   "Carrier_55_Carrier_Number_Echo" AT %QW3102 : Word;
   "Carrier_55_Carrier_Position_Echo" AT %QD3104 : DWord;
   "Carrier_55_Next_Carrier_Number" AT %QW3108 : Word;
   "Carrier_55_Next_Stop_Position" AT %QD3110 : DWord;
   "Carrier_55_Drive_Command_Speed" AT %QW3114 : Word;
   "Carrier_55_Duplicate_Carrier_Number" AT %QW3116 : Word;
   "Carrier_55_First_Duplicate_Carrier_Position" AT %QD3118 : DWord;
   "Carrier_55_Second_Duplicate_Carrier_Position" AT %QD3122 : DWord;
   "Carrier_55_CommandWord" AT %QW3126 : Word;
   "Carrier_55_Heartbeat" AT %Q3126.0 : Bool;
   "Carrier_55_Drive_Forward_Command" AT %Q3126.1 : Bool;
   "Carrier_55_Fault_Reset" AT %Q3126.2 : Bool;
   "Carrier_55_At_Command_Position" AT %Q3126.3 : Bool;
   "Carrier_55_Duplicate_Carrier_Fault" AT %Q3126.4 : Bool;
   "Carrier_55_Motion_On_Fault" AT %Q3126.5 : Bool;
   "Carrier_55_Motion_Off_Fault" AT %Q3126.6 : Bool;
   "Carrier_55_Carrier_Spacing_Fault" AT %Q3126.7 : Bool;
   "Carrier_56_Carrier_In_Zone" AT %QW3150 : Word;
   "Carrier_56_Carrier_Number_Echo" AT %QW3152 : Word;
   "Carrier_56_Carrier_Position_Echo" AT %QD3154 : DWord;
   "Carrier_56_Next_Carrier_Number" AT %QW3158 : Word;
   "Carrier_56_Next_Stop_Position" AT %QD3160 : DWord;
   "Carrier_56_Drive_Command_Speed" AT %QW3164 : Word;
   "Carrier_56_Duplicate_Carrier_Number" AT %QW3166 : Word;
   "Carrier_56_First_Duplicate_Carrier_Position" AT %QD3168 : DWord;
   "Carrier_56_Second_Duplicate_Carrier_Position" AT %QD3172 : DWord;
   "Carrier_56_CommandWord" AT %QW3176 : Word;
   "Carrier_56_Heartbeat" AT %Q3176.0 : Bool;
   "Carrier_56_Drive_Forward_Command" AT %Q3176.1 : Bool;
   "Carrier_56_Fault_Reset" AT %Q3176.2 : Bool;
   "Carrier_56_At_Command_Position" AT %Q3176.3 : Bool;
   "Carrier_56_Duplicate_Carrier_Fault" AT %Q3176.4 : Bool;
   "Carrier_56_Motion_On_Fault" AT %Q3176.5 : Bool;
   "Carrier_56_Motion_Off_Fault" AT %Q3176.6 : Bool;
   "Carrier_56_Carrier_Spacing_Fault" AT %Q3176.7 : Bool;
   "Carrier_57_Carrier_In_Zone" AT %QW3200 : Word;
   "Carrier_57_Carrier_Number_Echo" AT %QW3202 : Word;
   "Carrier_57_Carrier_Position_Echo" AT %QD3204 : DWord;
   "Carrier_57_Next_Carrier_Number" AT %QW3208 : Word;
   "Carrier_57_Next_Stop_Position" AT %QD3210 : DWord;
   "Carrier_57_Drive_Command_Speed" AT %QW3214 : Word;
   "Carrier_57_Duplicate_Carrier_Number" AT %QW3216 : Word;
   "Carrier_57_First_Duplicate_Carrier_Position" AT %QD3218 : DWord;
   "Carrier_57_Second_Duplicate_Carrier_Position" AT %QD3222 : DWord;
   "Carrier_57_CommandWord" AT %QW3226 : Word;
   "Carrier_57_Heartbeat" AT %Q3226.0 : Bool;
   "Carrier_57_Drive_Forward_Command" AT %Q3226.1 : Bool;
   "Carrier_57_Fault_Reset" AT %Q3226.2 : Bool;
   "Carrier_57_At_Command_Position" AT %Q3226.3 : Bool;
   "Carrier_57_Duplicate_Carrier_Fault" AT %Q3226.4 : Bool;
   "Carrier_57_Motion_On_Fault" AT %Q3226.5 : Bool;
   "Carrier_57_Motion_Off_Fault" AT %Q3226.6 : Bool;
   "Carrier_57_Carrier_Spacing_Fault" AT %Q3226.7 : Bool;
   "Carrier_58_Carrier_In_Zone" AT %QW3250 : Word;
   "Carrier_58_Carrier_Number_Echo" AT %QW3252 : Word;
   "Carrier_58_Carrier_Position_Echo" AT %QD3254 : DWord;
   "Carrier_58_Next_Carrier_Number" AT %QW3258 : Word;
   "Carrier_58_Next_Stop_Position" AT %QD3260 : DWord;
   "Carrier_58_Drive_Command_Speed" AT %QW3264 : Word;
   "Carrier_58_Duplicate_Carrier_Number" AT %QW3266 : Word;
   "Carrier_58_First_Duplicate_Carrier_Position" AT %QD3268 : DWord;
   "Carrier_58_Second_Duplicate_Carrier_Position" AT %QD3272 : DWord;
   "Carrier_58_CommandWord" AT %QW3276 : Word;
   "Carrier_58_Heartbeat" AT %Q3276.0 : Bool;
   "Carrier_58_Drive_Forward_Command" AT %Q3276.1 : Bool;
   "Carrier_58_Fault_Reset" AT %Q3276.2 : Bool;
   "Carrier_58_At_Command_Position" AT %Q3276.3 : Bool;
   "Carrier_58_Duplicate_Carrier_Fault" AT %Q3276.4 : Bool;
   "Carrier_58_Motion_On_Fault" AT %Q3276.5 : Bool;
   "Carrier_58_Motion_Off_Fault" AT %Q3276.6 : Bool;
   "Carrier_58_Carrier_Spacing_Fault" AT %Q3276.7 : Bool;
   "Carrier_59_Carrier_In_Zone" AT %QW3300 : Word;
   "Carrier_59_Carrier_Number_Echo" AT %QW3302 : Word;
   "Carrier_59_Carrier_Position_Echo" AT %QD3304 : DWord;
   "Carrier_59_Next_Carrier_Number" AT %QW3308 : Word;
   "Carrier_59_Next_Stop_Position" AT %QD3310 : DWord;
   "Carrier_59_Drive_Command_Speed" AT %QW3314 : Word;
   "Carrier_59_Duplicate_Carrier_Number" AT %QW3316 : Word;
   "Carrier_59_First_Duplicate_Carrier_Position" AT %QD3318 : DWord;
   "Carrier_59_Second_Duplicate_Carrier_Position" AT %QD3322 : DWord;
   "Carrier_59_CommandWord" AT %QW3326 : Word;
   "Carrier_59_Heartbeat" AT %Q3326.0 : Bool;
   "Carrier_59_Drive_Forward_Command" AT %Q3326.1 : Bool;
   "Carrier_59_Fault_Reset" AT %Q3326.2 : Bool;
   "Carrier_59_At_Command_Position" AT %Q3326.3 : Bool;
   "Carrier_59_Duplicate_Carrier_Fault" AT %Q3326.4 : Bool;
   "Carrier_59_Motion_On_Fault" AT %Q3326.5 : Bool;
   "Carrier_59_Motion_Off_Fault" AT %Q3326.6 : Bool;
   "Carrier_59_Carrier_Spacing_Fault" AT %Q3326.7 : Bool;
   "Carrier_60_Carrier_In_Zone" AT %QW3350 : Word;
   "Carrier_60_Carrier_Number_Echo" AT %QW3352 : Word;
   "Carrier_60_Carrier_Position_Echo" AT %QD3354 : DWord;
   "Carrier_60_Next_Carrier_Number" AT %QW3358 : Word;
   "Carrier_60_Next_Stop_Position" AT %QD3360 : DWord;
   "Carrier_60_Drive_Command_Speed" AT %QW3364 : Word;
   "Carrier_60_Duplicate_Carrier_Number" AT %QW3366 : Word;
   "Carrier_60_First_Duplicate_Carrier_Position" AT %QD3368 : DWord;
   "Carrier_60_Second_Duplicate_Carrier_Position" AT %QD3372 : DWord;
   "Carrier_60_CommandWord" AT %QW3376 : Word;
   "Carrier_60_Heartbeat" AT %Q3376.0 : Bool;
   "Carrier_60_Drive_Forward_Command" AT %Q3376.1 : Bool;
   "Carrier_60_Fault_Reset" AT %Q3376.2 : Bool;
   "Carrier_60_At_Command_Position" AT %Q3376.3 : Bool;
   "Carrier_60_Duplicate_Carrier_Fault" AT %Q3376.4 : Bool;
   "Carrier_60_Motion_On_Fault" AT %Q3376.5 : Bool;
   "Carrier_60_Motion_Off_Fault" AT %Q3376.6 : Bool;
   "Carrier_60_Carrier_Spacing_Fault" AT %Q3376.7 : Bool;
   "Carrier_61_Carrier_In_Zone" AT %QW3400 : Word;
   "Carrier_61_Carrier_Number_Echo" AT %QW3402 : Word;
   "Carrier_61_Carrier_Position_Echo" AT %QD3404 : DWord;
   "Carrier_61_Next_Carrier_Number" AT %QW3408 : Word;
   "Carrier_61_Next_Stop_Position" AT %QD3410 : DWord;
   "Carrier_61_Drive_Command_Speed" AT %QW3414 : Word;
   "Carrier_61_Duplicate_Carrier_Number" AT %QW3416 : Word;
   "Carrier_61_First_Duplicate_Carrier_Position" AT %QD3418 : DWord;
   "Carrier_61_Second_Duplicate_Carrier_Position" AT %QD3422 : DWord;
   "Carrier_61_CommandWord" AT %QW3426 : Word;
   "Carrier_61_Heartbeat" AT %Q3426.0 : Bool;
   "Carrier_61_Drive_Forward_Command" AT %Q3426.1 : Bool;
   "Carrier_61_Fault_Reset" AT %Q3426.2 : Bool;
   "Carrier_61_At_Command_Position" AT %Q3426.3 : Bool;
   "Carrier_61_Duplicate_Carrier_Fault" AT %Q3426.4 : Bool;
   "Carrier_61_Motion_On_Fault" AT %Q3426.5 : Bool;
   "Carrier_61_Motion_Off_Fault" AT %Q3426.6 : Bool;
   "Carrier_61_Carrier_Spacing_Fault" AT %Q3426.7 : Bool;
   "Carrier_62_Carrier_In_Zone" AT %QW3450 : Word;
   "Carrier_62_Carrier_Number_Echo" AT %QW3452 : Word;
   "Carrier_62_Carrier_Position_Echo" AT %QD3454 : DWord;
   "Carrier_62_Next_Carrier_Number" AT %QW3458 : Word;
   "Carrier_62_Next_Stop_Position" AT %QD3460 : DWord;
   "Carrier_62_Drive_Command_Speed" AT %QW3464 : Word;
   "Carrier_62_Duplicate_Carrier_Number" AT %QW3466 : Word;
   "Carrier_62_First_Duplicate_Carrier_Position" AT %QD3468 : DWord;
   "Carrier_62_Second_Duplicate_Carrier_Position" AT %QD3472 : DWord;
   "Carrier_62_CommandWord" AT %QW3476 : Word;
   "Carrier_62_Heartbeat" AT %Q3476.0 : Bool;
   "Carrier_62_Drive_Forward_Command" AT %Q3476.1 : Bool;
   "Carrier_62_Fault_Reset" AT %Q3476.2 : Bool;
   "Carrier_62_At_Command_Position" AT %Q3476.3 : Bool;
   "Carrier_62_Duplicate_Carrier_Fault" AT %Q3476.4 : Bool;
   "Carrier_62_Motion_On_Fault" AT %Q3476.5 : Bool;
   "Carrier_62_Motion_Off_Fault" AT %Q3476.6 : Bool;
   "Carrier_62_Carrier_Spacing_Fault" AT %Q3476.7 : Bool;
   "Carrier_63_Carrier_In_Zone" AT %QW3500 : Word;
   "Carrier_63_Carrier_Number_Echo" AT %QW3502 : Word;
   "Carrier_63_Carrier_Position_Echo" AT %QD3504 : DWord;
   "Carrier_63_Next_Carrier_Number" AT %QW3508 : Word;
   "Carrier_63_Next_Stop_Position" AT %QD3510 : DWord;
   "Carrier_63_Drive_Command_Speed" AT %QW3514 : Word;
   "Carrier_63_Duplicate_Carrier_Number" AT %QW3516 : Word;
   "Carrier_63_First_Duplicate_Carrier_Position" AT %QD3518 : DWord;
   "Carrier_63_Second_Duplicate_Carrier_Position" AT %QD3522 : DWord;
   "Carrier_63_CommandWord" AT %QW3526 : Word;
   "Carrier_63_Heartbeat" AT %Q3526.0 : Bool;
   "Carrier_63_Drive_Forward_Command" AT %Q3526.1 : Bool;
   "Carrier_63_Fault_Reset" AT %Q3526.2 : Bool;
   "Carrier_63_At_Command_Position" AT %Q3526.3 : Bool;
   "Carrier_63_Duplicate_Carrier_Fault" AT %Q3526.4 : Bool;
   "Carrier_63_Motion_On_Fault" AT %Q3526.5 : Bool;
   "Carrier_63_Motion_Off_Fault" AT %Q3526.6 : Bool;
   "Carrier_63_Carrier_Spacing_Fault" AT %Q3526.7 : Bool;
   "Carrier_64_Carrier_In_Zone" AT %QW3550 : Word;
   "Carrier_64_Carrier_Number_Echo" AT %QW3552 : Word;
   "Carrier_64_Carrier_Position_Echo" AT %QD3554 : DWord;
   "Carrier_64_Next_Carrier_Number" AT %QW3558 : Word;
   "Carrier_64_Next_Stop_Position" AT %QD3560 : DWord;
   "Carrier_64_Drive_Command_Speed" AT %QW3564 : Word;
   "Carrier_64_Duplicate_Carrier_Number" AT %QW3566 : Word;
   "Carrier_64_First_Duplicate_Carrier_Position" AT %QD3568 : DWord;
   "Carrier_64_Second_Duplicate_Carrier_Position" AT %QD3572 : DWord;
   "Carrier_64_CommandWord" AT %QW3576 : Word;
   "Carrier_64_Heartbeat" AT %Q3576.0 : Bool;
   "Carrier_64_Drive_Forward_Command" AT %Q3576.1 : Bool;
   "Carrier_64_Fault_Reset" AT %Q3576.2 : Bool;
   "Carrier_64_At_Command_Position" AT %Q3576.3 : Bool;
   "Carrier_64_Duplicate_Carrier_Fault" AT %Q3576.4 : Bool;
   "Carrier_64_Motion_On_Fault" AT %Q3576.5 : Bool;
   "Carrier_64_Motion_Off_Fault" AT %Q3576.6 : Bool;
   "Carrier_64_Carrier_Spacing_Fault" AT %Q3576.7 : Bool;
   "Carrier_65_Carrier_In_Zone" AT %QW3600 : Word;
   "Carrier_65_Carrier_Number_Echo" AT %QW3602 : Word;
   "Carrier_65_Carrier_Position_Echo" AT %QD3604 : DWord;
   "Carrier_65_Next_Carrier_Number" AT %QW3608 : Word;
   "Carrier_65_Next_Stop_Position" AT %QD3610 : DWord;
   "Carrier_65_Drive_Command_Speed" AT %QW3614 : Word;
   "Carrier_65_Duplicate_Carrier_Number" AT %QW3616 : Word;
   "Carrier_65_First_Duplicate_Carrier_Position" AT %QD3618 : DWord;
   "Carrier_65_Second_Duplicate_Carrier_Position" AT %QD3622 : DWord;
   "Carrier_65_CommandWord" AT %QW3626 : Word;
   "Carrier_65_Heartbeat" AT %Q3626.0 : Bool;
   "Carrier_65_Drive_Forward_Command" AT %Q3626.1 : Bool;
   "Carrier_65_Fault_Reset" AT %Q3626.2 : Bool;
   "Carrier_65_At_Command_Position" AT %Q3626.3 : Bool;
   "Carrier_65_Duplicate_Carrier_Fault" AT %Q3626.4 : Bool;
   "Carrier_65_Motion_On_Fault" AT %Q3626.5 : Bool;
   "Carrier_65_Motion_Off_Fault" AT %Q3626.6 : Bool;
   "Carrier_65_Carrier_Spacing_Fault" AT %Q3626.7 : Bool;
   "Carrier_66_Carrier_In_Zone" AT %QW3650 : Word;
   "Carrier_66_Carrier_Number_Echo" AT %QW3652 : Word;
   "Carrier_66_Carrier_Position_Echo" AT %QD3654 : DWord;
   "Carrier_66_Next_Carrier_Number" AT %QW3658 : Word;
   "Carrier_66_Next_Stop_Position" AT %QD3660 : DWord;
   "Carrier_66_Drive_Command_Speed" AT %QW3664 : Word;
   "Carrier_66_Duplicate_Carrier_Number" AT %QW3666 : Word;
   "Carrier_66_First_Duplicate_Carrier_Position" AT %QD3668 : DWord;
   "Carrier_66_Second_Duplicate_Carrier_Position" AT %QD3672 : DWord;
   "Carrier_66_CommandWord" AT %QW3676 : Word;
   "Carrier_66_Heartbeat" AT %Q3676.0 : Bool;
   "Carrier_66_Drive_Forward_Command" AT %Q3676.1 : Bool;
   "Carrier_66_Fault_Reset" AT %Q3676.2 : Bool;
   "Carrier_66_At_Command_Position" AT %Q3676.3 : Bool;
   "Carrier_66_Duplicate_Carrier_Fault" AT %Q3676.4 : Bool;
   "Carrier_66_Motion_On_Fault" AT %Q3676.5 : Bool;
   "Carrier_66_Motion_Off_Fault" AT %Q3676.6 : Bool;
   "Carrier_66_Carrier_Spacing_Fault" AT %Q3676.7 : Bool;
   "Carrier_67_Carrier_In_Zone" AT %QW3700 : Word;
   "Carrier_67_Carrier_Number_Echo" AT %QW3702 : Word;
   "Carrier_67_Carrier_Position_Echo" AT %QD3704 : DWord;
   "Carrier_67_Next_Carrier_Number" AT %QW3708 : Word;
   "Carrier_67_Next_Stop_Position" AT %QD3710 : DWord;
   "Carrier_67_Drive_Command_Speed" AT %QW3714 : Word;
   "Carrier_67_Duplicate_Carrier_Number" AT %QW3716 : Word;
   "Carrier_67_First_Duplicate_Carrier_Position" AT %QD3718 : DWord;
   "Carrier_67_Second_Duplicate_Carrier_Position" AT %QD3722 : DWord;
   "Carrier_67_CommandWord" AT %QW3726 : Word;
   "Carrier_67_Heartbeat" AT %Q3726.0 : Bool;
   "Carrier_67_Drive_Forward_Command" AT %Q3726.1 : Bool;
   "Carrier_67_Fault_Reset" AT %Q3726.2 : Bool;
   "Carrier_67_At_Command_Position" AT %Q3726.3 : Bool;
   "Carrier_67_Duplicate_Carrier_Fault" AT %Q3726.4 : Bool;
   "Carrier_67_Motion_On_Fault" AT %Q3726.5 : Bool;
   "Carrier_67_Motion_Off_Fault" AT %Q3726.6 : Bool;
   "Carrier_67_Carrier_Spacing_Fault" AT %Q3726.7 : Bool;
   "Carrier_68_Carrier_In_Zone" AT %QW3750 : Word;
   "Carrier_68_Carrier_Number_Echo" AT %QW3752 : Word;
   "Carrier_68_Carrier_Position_Echo" AT %QD3754 : DWord;
   "Carrier_68_Next_Carrier_Number" AT %QW3758 : Word;
   "Carrier_68_Next_Stop_Position" AT %QD3760 : DWord;
   "Carrier_68_Drive_Command_Speed" AT %QW3764 : Word;
   "Carrier_68_Duplicate_Carrier_Number" AT %QW3766 : Word;
   "Carrier_68_First_Duplicate_Carrier_Position" AT %QD3768 : DWord;
   "Carrier_68_Second_Duplicate_Carrier_Position" AT %QD3772 : DWord;
   "Carrier_68_CommandWord" AT %QW3776 : Word;
   "Carrier_68_Heartbeat" AT %Q3776.0 : Bool;
   "Carrier_68_Drive_Forward_Command" AT %Q3776.1 : Bool;
   "Carrier_68_Fault_Reset" AT %Q3776.2 : Bool;
   "Carrier_68_At_Command_Position" AT %Q3776.3 : Bool;
   "Carrier_68_Duplicate_Carrier_Fault" AT %Q3776.4 : Bool;
   "Carrier_68_Motion_On_Fault" AT %Q3776.5 : Bool;
   "Carrier_68_Motion_Off_Fault" AT %Q3776.6 : Bool;
   "Carrier_68_Carrier_Spacing_Fault" AT %Q3776.7 : Bool;
   "Carrier_69_Carrier_In_Zone" AT %QW3800 : Word;
   "Carrier_69_Carrier_Number_Echo" AT %QW3802 : Word;
   "Carrier_69_Carrier_Position_Echo" AT %QD3804 : DWord;
   "Carrier_69_Next_Carrier_Number" AT %QW3808 : Word;
   "Carrier_69_Next_Stop_Position" AT %QD3810 : DWord;
   "Carrier_69_Drive_Command_Speed" AT %QW3814 : Word;
   "Carrier_69_Duplicate_Carrier_Number" AT %QW3816 : Word;
   "Carrier_69_First_Duplicate_Carrier_Position" AT %QD3818 : DWord;
   "Carrier_69_Second_Duplicate_Carrier_Position" AT %QD3822 : DWord;
   "Carrier_69_CommandWord" AT %QW3826 : Word;
   "Carrier_69_Heartbeat" AT %Q3826.0 : Bool;
   "Carrier_69_Drive_Forward_Command" AT %Q3826.1 : Bool;
   "Carrier_69_Fault_Reset" AT %Q3826.2 : Bool;
   "Carrier_69_At_Command_Position" AT %Q3826.3 : Bool;
   "Carrier_69_Duplicate_Carrier_Fault" AT %Q3826.4 : Bool;
   "Carrier_69_Motion_On_Fault" AT %Q3826.5 : Bool;
   "Carrier_69_Motion_Off_Fault" AT %Q3826.6 : Bool;
   "Carrier_69_Carrier_Spacing_Fault" AT %Q3826.7 : Bool;
   "Carrier_70_Carrier_In_Zone" AT %QW3850 : Word;
   "Carrier_70_Carrier_Number_Echo" AT %QW3852 : Word;
   "Carrier_70_Carrier_Position_Echo" AT %QD3854 : DWord;
   "Carrier_70_Next_Carrier_Number" AT %QW3858 : Word;
   "Carrier_70_Next_Stop_Position" AT %QD3860 : DWord;
   "Carrier_70_Drive_Command_Speed" AT %QW3864 : Word;
   "Carrier_70_Duplicate_Carrier_Number" AT %QW3866 : Word;
   "Carrier_70_First_Duplicate_Carrier_Position" AT %QD3868 : DWord;
   "Carrier_70_Second_Duplicate_Carrier_Position" AT %QD3872 : DWord;
   "Carrier_70_CommandWord" AT %QW3876 : Word;
   "Carrier_70_Heartbeat" AT %Q3876.0 : Bool;
   "Carrier_70_Drive_Forward_Command" AT %Q3876.1 : Bool;
   "Carrier_70_Fault_Reset" AT %Q3876.2 : Bool;
   "Carrier_70_At_Command_Position" AT %Q3876.3 : Bool;
   "Carrier_70_Duplicate_Carrier_Fault" AT %Q3876.4 : Bool;
   "Carrier_70_Motion_On_Fault" AT %Q3876.5 : Bool;
   "Carrier_70_Motion_Off_Fault" AT %Q3876.6 : Bool;
   "Carrier_70_Carrier_Spacing_Fault" AT %Q3876.7 : Bool;
   "Carrier_71_Carrier_In_Zone" AT %QW3900 : Word;
   "Carrier_71_Carrier_Number_Echo" AT %QW3902 : Word;
   "Carrier_71_Carrier_Position_Echo" AT %QD3904 : DWord;
   "Carrier_71_Next_Carrier_Number" AT %QW3908 : Word;
   "Carrier_71_Next_Stop_Position" AT %QD3910 : DWord;
   "Carrier_71_Drive_Command_Speed" AT %QW3914 : Word;
   "Carrier_71_Duplicate_Carrier_Number" AT %QW3916 : Word;
   "Carrier_71_First_Duplicate_Carrier_Position" AT %QD3918 : DWord;
   "Carrier_71_Second_Duplicate_Carrier_Position" AT %QD3922 : DWord;
   "Carrier_71_CommandWord" AT %QW3926 : Word;
   "Carrier_71_Heartbeat" AT %Q3926.0 : Bool;
   "Carrier_71_Drive_Forward_Command" AT %Q3926.1 : Bool;
   "Carrier_71_Fault_Reset" AT %Q3926.2 : Bool;
   "Carrier_71_At_Command_Position" AT %Q3926.3 : Bool;
   "Carrier_71_Duplicate_Carrier_Fault" AT %Q3926.4 : Bool;
   "Carrier_71_Motion_On_Fault" AT %Q3926.5 : Bool;
   "Carrier_71_Motion_Off_Fault" AT %Q3926.6 : Bool;
   "Carrier_71_Carrier_Spacing_Fault" AT %Q3926.7 : Bool;
   "Carrier_72_Carrier_In_Zone" AT %QW3950 : Word;
   "Carrier_72_Carrier_Number_Echo" AT %QW3952 : Word;
   "Carrier_72_Carrier_Position_Echo" AT %QD3954 : DWord;
   "Carrier_72_Next_Carrier_Number" AT %QW3958 : Word;
   "Carrier_72_Next_Stop_Position" AT %QD3960 : DWord;
   "Carrier_72_Drive_Command_Speed" AT %QW3964 : Word;
   "Carrier_72_Duplicate_Carrier_Number" AT %QW3966 : Word;
   "Carrier_72_First_Duplicate_Carrier_Position" AT %QD3968 : DWord;
   "Carrier_72_Second_Duplicate_Carrier_Position" AT %QD3972 : DWord;
   "Carrier_72_CommandWord" AT %QW3976 : Word;
   "Carrier_72_Heartbeat" AT %Q3976.0 : Bool;
   "Carrier_72_Drive_Forward_Command" AT %Q3976.1 : Bool;
   "Carrier_72_Fault_Reset" AT %Q3976.2 : Bool;
   "Carrier_72_At_Command_Position" AT %Q3976.3 : Bool;
   "Carrier_72_Duplicate_Carrier_Fault" AT %Q3976.4 : Bool;
   "Carrier_72_Motion_On_Fault" AT %Q3976.5 : Bool;
   "Carrier_72_Motion_Off_Fault" AT %Q3976.6 : Bool;
   "Carrier_72_Carrier_Spacing_Fault" AT %Q3976.7 : Bool;
   "Carrier_73_Carrier_In_Zone" AT %QW4000 : Word;
   "Carrier_73_Carrier_Number_Echo" AT %QW4002 : Word;
   "Carrier_73_Carrier_Position_Echo" AT %QD4004 : DWord;
   "Carrier_73_Next_Carrier_Number" AT %QW4008 : Word;
   "Carrier_73_Next_Stop_Position" AT %QD4010 : DWord;
   "Carrier_73_Drive_Command_Speed" AT %QW4014 : Word;
   "Carrier_73_Duplicate_Carrier_Number" AT %QW4016 : Word;
   "Carrier_73_First_Duplicate_Carrier_Position" AT %QD4018 : DWord;
   "Carrier_73_Second_Duplicate_Carrier_Position" AT %QD4022 : DWord;
   "Carrier_73_CommandWord" AT %QW4026 : Word;
   "Carrier_73_Heartbeat" AT %Q4026.0 : Bool;
   "Carrier_73_Drive_Forward_Command" AT %Q4026.1 : Bool;
   "Carrier_73_Fault_Reset" AT %Q4026.2 : Bool;
   "Carrier_73_At_Command_Position" AT %Q4026.3 : Bool;
   "Carrier_73_Duplicate_Carrier_Fault" AT %Q4026.4 : Bool;
   "Carrier_73_Motion_On_Fault" AT %Q4026.5 : Bool;
   "Carrier_73_Motion_Off_Fault" AT %Q4026.6 : Bool;
   "Carrier_73_Carrier_Spacing_Fault" AT %Q4026.7 : Bool;
   "Carrier_74_Carrier_In_Zone" AT %QW4050 : Word;
   "Carrier_74_Carrier_Number_Echo" AT %QW4052 : Word;
   "Carrier_74_Carrier_Position_Echo" AT %QD4054 : DWord;
   "Carrier_74_Next_Carrier_Number" AT %QW4058 : Word;
   "Carrier_74_Next_Stop_Position" AT %QD4060 : DWord;
   "Carrier_74_Drive_Command_Speed" AT %QW4064 : Word;
   "Carrier_74_Duplicate_Carrier_Number" AT %QW4066 : Word;
   "Carrier_74_First_Duplicate_Carrier_Position" AT %QD4068 : DWord;
   "Carrier_74_Second_Duplicate_Carrier_Position" AT %QD4072 : DWord;
   "Carrier_74_CommandWord" AT %QW4076 : Word;
   "Carrier_74_Heartbeat" AT %Q4076.0 : Bool;
   "Carrier_74_Drive_Forward_Command" AT %Q4076.1 : Bool;
   "Carrier_74_Fault_Reset" AT %Q4076.2 : Bool;
   "Carrier_74_At_Command_Position" AT %Q4076.3 : Bool;
   "Carrier_74_Duplicate_Carrier_Fault" AT %Q4076.4 : Bool;
   "Carrier_74_Motion_On_Fault" AT %Q4076.5 : Bool;
   "Carrier_74_Motion_Off_Fault" AT %Q4076.6 : Bool;
   "Carrier_74_Carrier_Spacing_Fault" AT %Q4076.7 : Bool;
   "Carrier_75_Carrier_In_Zone" AT %QW4100 : Word;
   "Carrier_75_Carrier_Number_Echo" AT %QW4102 : Word;
   "Carrier_75_Carrier_Position_Echo" AT %QD4104 : DWord;
   "Carrier_75_Next_Carrier_Number" AT %QW4108 : Word;
   "Carrier_75_Next_Stop_Position" AT %QD4110 : DWord;
   "Carrier_75_Drive_Command_Speed" AT %QW4114 : Word;
   "Carrier_75_Duplicate_Carrier_Number" AT %QW4116 : Word;
   "Carrier_75_First_Duplicate_Carrier_Position" AT %QD4118 : DWord;
   "Carrier_75_Second_Duplicate_Carrier_Position" AT %QD4122 : DWord;
   "Carrier_75_CommandWord" AT %QW4126 : Word;
   "Carrier_75_Heartbeat" AT %Q4126.0 : Bool;
   "Carrier_75_Drive_Forward_Command" AT %Q4126.1 : Bool;
   "Carrier_75_Fault_Reset" AT %Q4126.2 : Bool;
   "Carrier_75_At_Command_Position" AT %Q4126.3 : Bool;
   "Carrier_75_Duplicate_Carrier_Fault" AT %Q4126.4 : Bool;
   "Carrier_75_Motion_On_Fault" AT %Q4126.5 : Bool;
   "Carrier_75_Motion_Off_Fault" AT %Q4126.6 : Bool;
   "Carrier_75_Carrier_Spacing_Fault" AT %Q4126.7 : Bool;
   "Carrier_76_Carrier_In_Zone" AT %QW4150 : Word;
   "Carrier_76_Carrier_Number_Echo" AT %QW4152 : Word;
   "Carrier_76_Carrier_Position_Echo" AT %QD4154 : DWord;
   "Carrier_76_Next_Carrier_Number" AT %QW4158 : Word;
   "Carrier_76_Next_Stop_Position" AT %QD4160 : DWord;
   "Carrier_76_Drive_Command_Speed" AT %QW4164 : Word;
   "Carrier_76_Duplicate_Carrier_Number" AT %QW4166 : Word;
   "Carrier_76_First_Duplicate_Carrier_Position" AT %QD4168 : DWord;
   "Carrier_76_Second_Duplicate_Carrier_Position" AT %QD4172 : DWord;
   "Carrier_76_CommandWord" AT %QW4176 : Word;
   "Carrier_76_Heartbeat" AT %Q4176.0 : Bool;
   "Carrier_76_Drive_Forward_Command" AT %Q4176.1 : Bool;
   "Carrier_76_Fault_Reset" AT %Q4176.2 : Bool;
   "Carrier_76_At_Command_Position" AT %Q4176.3 : Bool;
   "Carrier_76_Duplicate_Carrier_Fault" AT %Q4176.4 : Bool;
   "Carrier_76_Motion_On_Fault" AT %Q4176.5 : Bool;
   "Carrier_76_Motion_Off_Fault" AT %Q4176.6 : Bool;
   "Carrier_76_Carrier_Spacing_Fault" AT %Q4176.7 : Bool;
   "Carrier_77_Carrier_In_Zone" AT %QW4200 : Word;
   "Carrier_77_Carrier_Number_Echo" AT %QW4202 : Word;
   "Carrier_77_Carrier_Position_Echo" AT %QD4204 : DWord;
   "Carrier_77_Next_Carrier_Number" AT %QW4208 : Word;
   "Carrier_77_Next_Stop_Position" AT %QD4210 : DWord;
   "Carrier_77_Drive_Command_Speed" AT %QW4214 : Word;
   "Carrier_77_Duplicate_Carrier_Number" AT %QW4216 : Word;
   "Carrier_77_First_Duplicate_Carrier_Position" AT %QD4218 : DWord;
   "Carrier_77_Second_Duplicate_Carrier_Position" AT %QD4222 : DWord;
   "Carrier_77_CommandWord" AT %QW4226 : Word;
   "Carrier_77_Heartbeat" AT %Q4226.0 : Bool;
   "Carrier_77_Drive_Forward_Command" AT %Q4226.1 : Bool;
   "Carrier_77_Fault_Reset" AT %Q4226.2 : Bool;
   "Carrier_77_At_Command_Position" AT %Q4226.3 : Bool;
   "Carrier_77_Duplicate_Carrier_Fault" AT %Q4226.4 : Bool;
   "Carrier_77_Motion_On_Fault" AT %Q4226.5 : Bool;
   "Carrier_77_Motion_Off_Fault" AT %Q4226.6 : Bool;
   "Carrier_77_Carrier_Spacing_Fault" AT %Q4226.7 : Bool;
   "Carrier_78_Carrier_In_Zone" AT %QW4250 : Word;
   "Carrier_78_Carrier_Number_Echo" AT %QW4252 : Word;
   "Carrier_78_Carrier_Position_Echo" AT %QD4254 : DWord;
   "Carrier_78_Next_Carrier_Number" AT %QW4258 : Word;
   "Carrier_78_Next_Stop_Position" AT %QD4260 : DWord;
   "Carrier_78_Drive_Command_Speed" AT %QW4264 : Word;
   "Carrier_78_Duplicate_Carrier_Number" AT %QW4266 : Word;
   "Carrier_78_First_Duplicate_Carrier_Position" AT %QD4268 : DWord;
   "Carrier_78_Second_Duplicate_Carrier_Position" AT %QD4272 : DWord;
   "Carrier_78_CommandWord" AT %QW4276 : Word;
   "Carrier_78_Heartbeat" AT %Q4276.0 : Bool;
   "Carrier_78_Drive_Forward_Command" AT %Q4276.1 : Bool;
   "Carrier_78_Fault_Reset" AT %Q4276.2 : Bool;
   "Carrier_78_At_Command_Position" AT %Q4276.3 : Bool;
   "Carrier_78_Duplicate_Carrier_Fault" AT %Q4276.4 : Bool;
   "Carrier_78_Motion_On_Fault" AT %Q4276.5 : Bool;
   "Carrier_78_Motion_Off_Fault" AT %Q4276.6 : Bool;
   "Carrier_78_Carrier_Spacing_Fault" AT %Q4276.7 : Bool;
   "Carrier_79_Carrier_In_Zone" AT %QW4300 : Word;
   "Carrier_79_Carrier_Number_Echo" AT %QW4302 : Word;
   "Carrier_79_Carrier_Position_Echo" AT %QD4304 : DWord;
   "Carrier_79_Next_Carrier_Number" AT %QW4308 : Word;
   "Carrier_79_Next_Stop_Position" AT %QD4310 : DWord;
   "Carrier_79_Drive_Command_Speed" AT %QW4314 : Word;
   "Carrier_79_Duplicate_Carrier_Number" AT %QW4316 : Word;
   "Carrier_79_First_Duplicate_Carrier_Position" AT %QD4318 : DWord;
   "Carrier_79_Second_Duplicate_Carrier_Position" AT %QD4322 : DWord;
   "Carrier_79_CommandWord" AT %QW4326 : Word;
   "Carrier_79_Heartbeat" AT %Q4326.0 : Bool;
   "Carrier_79_Drive_Forward_Command" AT %Q4326.1 : Bool;
   "Carrier_79_Fault_Reset" AT %Q4326.2 : Bool;
   "Carrier_79_At_Command_Position" AT %Q4326.3 : Bool;
   "Carrier_79_Duplicate_Carrier_Fault" AT %Q4326.4 : Bool;
   "Carrier_79_Motion_On_Fault" AT %Q4326.5 : Bool;
   "Carrier_79_Motion_Off_Fault" AT %Q4326.6 : Bool;
   "Carrier_79_Carrier_Spacing_Fault" AT %Q4326.7 : Bool;
   "Carrier_80_Carrier_In_Zone" AT %QW4350 : Word;
   "Carrier_80_Carrier_Number_Echo" AT %QW4352 : Word;
   "Carrier_80_Carrier_Position_Echo" AT %QD4354 : DWord;
   "Carrier_80_Next_Carrier_Number" AT %QW4358 : Word;
   "Carrier_80_Next_Stop_Position" AT %QD4360 : DWord;
   "Carrier_80_Drive_Command_Speed" AT %QW4364 : Word;
   "Carrier_80_Duplicate_Carrier_Number" AT %QW4366 : Word;
   "Carrier_80_First_Duplicate_Carrier_Position" AT %QD4368 : DWord;
   "Carrier_80_Second_Duplicate_Carrier_Position" AT %QD4372 : DWord;
   "Carrier_80_CommandWord" AT %QW4376 : Word;
   "Carrier_80_Heartbeat" AT %Q4376.0 : Bool;
   "Carrier_80_Drive_Forward_Command" AT %Q4376.1 : Bool;
   "Carrier_80_Fault_Reset" AT %Q4376.2 : Bool;
   "Carrier_80_At_Command_Position" AT %Q4376.3 : Bool;
   "Carrier_80_Duplicate_Carrier_Fault" AT %Q4376.4 : Bool;
   "Carrier_80_Motion_On_Fault" AT %Q4376.5 : Bool;
   "Carrier_80_Motion_Off_Fault" AT %Q4376.6 : Bool;
   "Carrier_80_Carrier_Spacing_Fault" AT %Q4376.7 : Bool;
   "Carrier_81_Carrier_In_Zone" AT %QW4400 : Word;
   "Carrier_81_Carrier_Number_Echo" AT %QW4402 : Word;
   "Carrier_81_Carrier_Position_Echo" AT %QD4404 : DWord;
   "Carrier_81_Next_Carrier_Number" AT %QW4408 : Word;
   "Carrier_81_Next_Stop_Position" AT %QD4410 : DWord;
   "Carrier_81_Drive_Command_Speed" AT %QW4414 : Word;
   "Carrier_81_Duplicate_Carrier_Number" AT %QW4416 : Word;
   "Carrier_81_First_Duplicate_Carrier_Position" AT %QD4418 : DWord;
   "Carrier_81_Second_Duplicate_Carrier_Position" AT %QD4422 : DWord;
   "Carrier_81_CommandWord" AT %QW4426 : Word;
   "Carrier_81_Heartbeat" AT %Q4426.0 : Bool;
   "Carrier_81_Drive_Forward_Command" AT %Q4426.1 : Bool;
   "Carrier_81_Fault_Reset" AT %Q4426.2 : Bool;
   "Carrier_81_At_Command_Position" AT %Q4426.3 : Bool;
   "Carrier_81_Duplicate_Carrier_Fault" AT %Q4426.4 : Bool;
   "Carrier_81_Motion_On_Fault" AT %Q4426.5 : Bool;
   "Carrier_81_Motion_Off_Fault" AT %Q4426.6 : Bool;
   "Carrier_81_Carrier_Spacing_Fault" AT %Q4426.7 : Bool;
   "Carrier_82_Carrier_In_Zone" AT %QW4450 : Word;
   "Carrier_82_Carrier_Number_Echo" AT %QW4452 : Word;
   "Carrier_82_Carrier_Position_Echo" AT %QD4454 : DWord;
   "Carrier_82_Next_Carrier_Number" AT %QW4458 : Word;
   "Carrier_82_Next_Stop_Position" AT %QD4460 : DWord;
   "Carrier_82_Drive_Command_Speed" AT %QW4464 : Word;
   "Carrier_82_Duplicate_Carrier_Number" AT %QW4466 : Word;
   "Carrier_82_First_Duplicate_Carrier_Position" AT %QD4468 : DWord;
   "Carrier_82_Second_Duplicate_Carrier_Position" AT %QD4472 : DWord;
   "Carrier_82_CommandWord" AT %QW4476 : Word;
   "Carrier_82_Heartbeat" AT %Q4476.0 : Bool;
   "Carrier_82_Drive_Forward_Command" AT %Q4476.1 : Bool;
   "Carrier_82_Fault_Reset" AT %Q4476.2 : Bool;
   "Carrier_82_At_Command_Position" AT %Q4476.3 : Bool;
   "Carrier_82_Duplicate_Carrier_Fault" AT %Q4476.4 : Bool;
   "Carrier_82_Motion_On_Fault" AT %Q4476.5 : Bool;
   "Carrier_82_Motion_Off_Fault" AT %Q4476.6 : Bool;
   "Carrier_82_Carrier_Spacing_Fault" AT %Q4476.7 : Bool;
END_VAR

VAR_GLOBAL   // PLC tag table "GW_EMS01_TO_SDC_TagTable"
   "EMS01_SDC_Stop1_Control" AT %IW10000 : Word;
   "EMS01_SDC_Stop2_Control" AT %IW10002 : Word;
   "EMS01_SDC_Stop3_Control" AT %IW10004 : Word;
   "EMS01_SDC_Stop4_Control" AT %IW10006 : Word;
   "EMS01_SDC_Stop5_Control" AT %IW10008 : Word;
   "EMS01_SDC_Stop6_Control" AT %IW10010 : Word;
   "EMS01_SDC_Stop7_Control" AT %IW10012 : Word;
   "EMS01_SDC_Stop8_Control" AT %IW10014 : Word;
   "EMS01_SDC_Stop9_Control" AT %IW10016 : Word;
   "EMS01_SDC_Stop10_Control" AT %IW10018 : Word;
   "EMS01_SDC_Stop11_Control" AT %IW10020 : Word;
   "EMS01_SDC_Stop12_Control" AT %IW10022 : Word;
   "EMS01_SDC_Stop13_Control" AT %IW10024 : Word;
   "EMS01_SDC_Stop14_Control" AT %IW10026 : Word;
   "EMS01_SDC_Stop15_Control" AT %IW10028 : Word;
   "EMS01_SDC_Stop16_Control" AT %IW10030 : Word;
   "EMS01_SDC_Stop17_Control" AT %IW10032 : Word;
   "EMS01_SDC_Stop18_Control" AT %IW10034 : Word;
   "EMS01_SDC_Stop19_Control" AT %IW10036 : Word;
   "EMS01_SDC_Stop20_Control" AT %IW10038 : Word;
   "EMS01_SDC_Stop21_Control" AT %IW10040 : Word;
   "EMS01_SDC_Stop22_Control" AT %IW10042 : Word;
   "EMS01_SDC_Stop23_Control" AT %IW10044 : Word;
   "EMS01_SDC_Stop24_Control" AT %IW10046 : Word;
   "EMS01_SDC_Stop25_Control" AT %IW10048 : Word;
   "EMS01_SDC_Stop26_Control" AT %IW10050 : Word;
   "EMS01_SDC_Stop27_Control" AT %IW10052 : Word;
   "EMS01_SDC_Stop28_Control" AT %IW10054 : Word;
   "EMS01_SDC_Stop29_Control" AT %IW10056 : Word;
   "EMS01_SDC_Stop30_Control" AT %IW10058 : Word;
   "EMS01_SDC_Stop31_Control" AT %IW10060 : Word;
   "EMS01_SDC_Stop32_Control" AT %IW10062 : Word;
   "EMS01_SDC_Stop33_Control" AT %IW10064 : Word;
   "EMS01_SDC_Stop34_Control" AT %IW10066 : Word;
   "EMS01_SDC_Stop35_Control" AT %IW10068 : Word;
   "EMS01_SDC_Stop36_Control" AT %IW10070 : Word;
   "EMS01_SDC_Stop37_Control" AT %IW10072 : Word;
   "EMS01_SDC_Stop38_Control" AT %IW10074 : Word;
   "EMS01_SDC_Stop39_Control" AT %IW10076 : Word;
   "EMS01_SDC_Stop40_Control" AT %IW10078 : Word;
   "EMS01_SDC_Stop41_Control" AT %IW10080 : Word;
   "EMS01_SDC_Stop42_Control" AT %IW10082 : Word;
   "EMS01_SDC_Stop43_Control" AT %IW10084 : Word;
   "EMS01_SDC_Stop44_Control" AT %IW10086 : Word;
   "EMS01_SDC_Stop45_Control" AT %IW10088 : Word;
   "EMS01_SDC_Stop46_Control" AT %IW10090 : Word;
   "EMS01_SDC_Stop47_Control" AT %IW10092 : Word;
   "EMS01_SDC_Stop48_Control" AT %IW10094 : Word;
   "EMS01_SDC_Stop49_Control" AT %IW10096 : Word;
   "EMS01_SDC_Stop50_Control" AT %IW10098 : Word;
   "EMS01_SDC_Stop51_Control" AT %IW10100 : Word;
   "EMS01_SDC_Stop52_Control" AT %IW10102 : Word;
   "EMS01_SDC_Stop53_Control" AT %IW10104 : Word;
   "EMS01_SDC_Stop54_Control" AT %IW10106 : Word;
   "EMS01_SDC_Stop55_Control" AT %IW10108 : Word;
   "EMS01_SDC_Stop56_Control" AT %IW10110 : Word;
   "EMS01_SDC_Stop57_Control" AT %IW10112 : Word;
   "EMS01_SDC_Stop58_Control" AT %IW10114 : Word;
   "EMS01_SDC_Stop59_Control" AT %IW10116 : Word;
   "EMS01_SDC_Stop60_Control" AT %IW10118 : Word;
   "EMS01_SDC_Stop61_Control" AT %IW10120 : Word;
   "EMS01_SDC_Stop62_Control" AT %IW10122 : Word;
   "EMS01_SDC_Stop63_Control" AT %IW10124 : Word;
   "EMS01_SDC_Stop64_Control" AT %IW10126 : Word;
   "EMS01_SDC_Stop65_Control" AT %IW10128 : Word;
   "EMS01_Status" AT %IW10150 : Word;
   "EMS01_MASTER_POWER_ON_ON_DELAY_" AT %I10150.0 : Bool;
   "EMS01_FAULT_RESET__PB_2406" AT %I10150.1 : Bool;
   "EMS01R1_MASTER_POWER_ON_ON_DELAY_" AT %I10150.2 : Bool;
   "EMS01R1_FAULT_RESET__PB_2406" AT %I10150.3 : Bool;
   "EMS01R2_MASTER_POWER_ON_ON_DELAY_" AT %I10150.4 : Bool;
   "EMS01R2_FAULT_RESET__PB_2406" AT %I10150.5 : Bool;
   "EMS01R3_MASTER_POWER_ON_ON_DELAY_" AT %I10150.6 : Bool;
   "EMS01R3_FAULT_RESET__PB_2406" AT %I10150.7 : Bool;
   "EMS01R4_MASTER_POWER_ON_ON_DELAY_" AT %I10151.0 : Bool;
   "EMS01R4_FAULT_RESET__PB_3206" AT %I10151.1 : Bool;
   "EMS01_Stop_#26__Set_To_Release" AT %I10151.2 : Bool;
   "EMS01_SpareBool1" AT %I10151.3 : Bool;
   "EMS01_SpareBool2" AT %I10151.4 : Bool;
   "EMS01_SpareBool3" AT %I10151.5 : Bool;
   "EMS01_SpareBool4" AT %I10151.6 : Bool;
   "EMS01_Heartbeat" AT %I10151.7 : Bool;
   "EMS01_SpareWord1" AT %IW10152 : Word;
   "EMS01_SpareWord2" AT %IW10154 : Word;
   "EMS01_CARRIER_SPEED_REF_160_ft_m" AT %IW10156 : Word;   // CARRIER_SPEED_REF_160_ft/m_=_-16768_130_ft/m_=_-25536_65_ft/m_=_20000_30_ft/m_=_9144
   "EMS01_PRODUCTION_SPEED_REF_(mm_min)__" AT %IW10158 : Word;
   "EMS01_PRODUCTION_SPEED_REF_(ft*10_min)__" AT %IW10160 : Word;
   "EMS01_PANELVIEW_#6_CARRIER_#_SELECTED_TO_BE_DELETED" AT %IW10174 : Word;
   "EMS01_SpareWord3" AT %IW10176 : Word;
   "EMS01_SpareWord4" AT %IW10178 : Word;
END_VAR

